(* Logix 5000 project; controller PLC_MCC1300_75F1 vendor 1 type 14 code 166 rev 32.11; software revision 32.04 *) (continued)
TYPE MAC_Conveyor_ALM :
STRUCT
   rgxStoppingFault : DINT[1];   // Generic stopping faults
   rgxFault : DINT[1];   // Generic faults
   rgxWarning : DINT[1];   // Generic warning
   rgxStoppingFault_M : DINT[2];   // Motor stopping faults
   rgxFault_M : DINT[2];   // Motor faults
   rgxWarning_M : DINT[2];   // Motor warning
   rgdFaultCode_M : DINT[2];   // Motor fault codes
END_STRUCT
END_TYPE

TYPE MAC_Conveyor_HMR :
STRUCT
   xSensorPresence1 : BOOL;   // Sensor presence 1 {x|x|x|x|O}
   xSensorPresence2 : BOOL;   // Sensor presence 2 {x|x|x|x|O}
   xSensorPresence3 : BOOL;   // Sensor presence 3 {x|x|x|x|O}
   xSensorPresence4 : BOOL;   // Sensor presence 4 {x|x|x|x|O}
   xSensorPresence5 : BOOL;   // Sensor presence 5 {x|x|x|x|O}
   xSensorPresence6 : BOOL;   // Sensor presence 6 {x|x|x|x|O}
   xHighPositionPopup1 : BOOL;   // High position popup {x|x|x|x|O}
   xLowPositionPopup1 : BOOL;   // Low position popup {x|x|x|x|O}
   xHighPositionPopup2 : BOOL;   // High position popup {x|x|x|x|O}
   xLowPositionPopup2 : BOOL;   // Low position popup {x|x|x|x|O}
   xHighPositionSquaring1 : BOOL;   // High position squaring {x|x|x|x|O}
   xLowPositionSquaring1 : BOOL;   // Low position squaring {x|x|x|x|O}
   xHighPositionSquaring2 : BOOL;   // High position squaring {x|x|x|x|O}
   xLowPositionSquaring2 : BOOL;   // Low position squaring {x|x|x|x|O}
   xCleaningEnabled : BOOL;   // Cleaning enabled {x|x|x|x|O}
   xWritingEnabled : BOOL;   // Writing enabled {x|x|x|x|O}
   xManualCommandEnabled : BOOL;   // Manual commands enabled {x|x|x|x|O}
   xVirtualDoorEnabled : BOOL;   // Virtual door enabled {x|x|x|x|O}
   xAuxFunctionEnabled : BOOL;   // Auxiliary function enabled {x|x|x|x|O}
   xIdPlatePresence : BOOL;   // Id plate presence {x|x|x|x|O}
   dState1 : DINT;   // State 1 (1=No anomaly, 3=Run, 7=Anomaly) {x|x|x|x|O}
   dState2 : DINT;   // State 2 (1=No anomaly, 3=Run, 7=Anomaly) {x|x|x|x|O}
   dState3 : DINT;   // State 3 (1=No anomaly, 3=Run, 7=Anomaly) {x|x|x|x|O}
   dState4 : DINT;   // State 4 (1=No anomaly, 3=Run, 7=Anomaly) {x|x|x|x|O}
   dStateSensor1 : DINT;   // State sensor 1 (1=No alarm, 7=Alarm) {x|x|x|x|O}
   dStateSensor2 : DINT;   // State sensor 2 (1=No alarm, 7=Alarm) {x|x|x|x|O}
   dStateSensor3 : DINT;   // State sensor 3(1=No alarm, 7=Alarm) {x|x|x|x|O}
   dStateSensor4 : DINT;   // State sensor 4(1=No alarm, 7=Alarm) {x|x|x|x|O}
   dStateSensor5 : DINT;   // State sensor 5(1=No alarm, 7=Alarm) {x|x|x|x|O}
   dStateSensor6 : DINT;   // State sensor 6(1=No alarm, 7=Alarm) {x|x|x|x|O}
   dErrorCode1 : DINT;   // Error code {x|x|x|x|O}
   dErrorCode2 : DINT;   // Error code {x|x|x|x|O}
   dErrorCode3 : DINT;   // Error code {x|x|x|x|O}
   dErrorCode4 : DINT;   // Error code {x|x|x|x|O}
   rgxMan : DINT;   // Manual commands {x|x|x|x|O}
END_STRUCT
END_TYPE

TYPE MAC_Conveyor_HMW :
STRUCT
   xLocalCleaningRequest : BOOL;   // Local cleaning request {x|x|x|x|O}
   xStopLocalCleaningRequest : BOOL;   // Stop local cleaning request {x|x|x|x|O}
   xEnableDisableManualCommand : BOOL;   // Enable/Disable manual commands {x|x|x|x|O}
   xSendDataToPLC : BOOL;   // Send plate data to PLC {x|x|x|x|O}
   xEnableDisableVirtualDoor : BOOL;   // Enable/Disable virtual door {x|x|x|x|O}
   xEnableDisableAuxFunction : BOOL;   // Enable/Disable auxiliary function {x|x|x|x|O}
   dParam_1_cmm : DINT;   // Auxiliary parameter 1 [mm/100] {mm/100|mm|x|x|O}
   dParam_2_cmm : DINT;   // Auxiliary parameter 2 [mm/100] {mm/100|mm|x|x|O}
   dParam_3_cmm : DINT;   // Auxiliary parameter 3 [mm/100] {mm/100|mm|x|x|O}
   dParam_4_cmm : DINT;   // Auxiliary parameter 4 [mm/100] {mm/100|mm|x|x|O}
   dParam_5_ms : DINT;   // Auxiliary parameter 5 [ms] {ms|ms|x|x|O}
   dParam_6_ms : DINT;   // Auxiliary parameter 6 [ms] {ms|ms|x|x|O}
   dParam_7_ms : DINT;   // Auxiliary parameter 7 [ms] {ms|ms|x|x|O}
   dParam_8_ms : DINT;   // Auxiliary parameter 8 [ms] {ms|ms|x|x|O}
   rgxMan : DINT;   // Manual commands {x|x|x|x|O}
END_STRUCT
END_TYPE

TYPE MAC_Conveyor_Single :
STRUCT
   ST_xInitialConditionOK : BOOL;   // Initial condition OK
   ST_xInitialConditionOK_BW : BOOL;   // Initial condition OK backward
   ST_xCleaningConditionOK : BOOL;   // Cleaning condition OK
   ST_xCleaningAccepted : BOOL;   // Cleaning accepted
   ST_xReqCleaning : BOOL;   // Request cleaning
   ST_xPlatePresence : BOOL;   // Plate presence memory
   ST_xPhasesInProgress : BOOL;   // Phases in progress
   ST_xCycleLoadUnload : BOOL;   // Cycle load/unload simultaneously
   ST_xStopMachineFault : BOOL;   // Stopped machine fault
   ST_xStopNextCycleFault : BOOL;   // Stop next cycle fault
   ST_xConditionOKStopCycle : BOOL;   // Condition OK for stop cycle
   ST_xOutputEnable : BOOL;   // Output enable
   ST_xMachineAlarm : BOOL;   // Machine alarm
   ST_xMachineWarning : BOOL;   // Machine warning
   ST_xIdPlatePresence : BOOL;   // Id plate presence
   ST_xFeedbackRotation : BOOL;   // Feedback rotation
   ST_xRampInProgress : BOOL;   // Ramp in progress
   ST_xAccInProgress : BOOL;   // Acceleration in progress
   ST_xDecInProgress : BOOL;   // Deceleration in progress
   ST_xWaitStopNextMachine : BOOL;   // Wait stop next machine
   ST_xWaitMachineStop : BOOL;   // Wait machine stop
   ST_xWaitReadyToMove : BOOL;   // Wait ready to move
   ST_xEnableControlError : BOOL;   // Enable control error
   ST_xManualMode : BOOL;   // Manual mode enabled
   ST_xPlateSynchronized : BOOL;   // Plate synchronized
   ST_xVirtualDoorEnabled : BOOL;   // Virtual door enabled
   ST_xDisableLoadUnloadOnStop : BOOL;   // Temporary disable of load/unload continuosly after a bit wait machine stop
   ST_xPlatePassageUpstream_FW : BOOL;   // Plate in passage upstream
   ST_xPlatePassageUpstream_BKW : BOOL;   // Plate in passage upstream
   ST_xPlatePassageDownstream_FW : BOOL;   // Plate in passage downstream
   ST_xPlatePassageDownstream_BKW : BOOL;   // Plate in passage downstream
   ST_xAxleReadyToMoveDelayed : BOOL;   // Axle ready to move delayed (NU)
   ST_xSafetyMovement : BOOL;   // Safety Mouvement
   ST_xReqDescent : BOOL;   // popup conveyor
   ST_xPhaseError : BOOL;   // Phase error, send lites to cullet
   ST_xAux1 : BOOL;   // ST Aux 1
   ST_xAux2 : BOOL;   // ST Aux 2
   ST_xAux3 : BOOL;   // ST Aux 3
   ST_xAux4 : BOOL;   // ST Aux 4
   OSR_xUnload : BOOL;   // OSR Unload
   OSR_xSynchroPhotocellHead : BOOL;   // OSR Synchronization photocell head
   OSR_xSynchroPhotocellTail : BOOL;   // OSR Synchronization photocell tail
   OSR_xPosReq : BOOL;   // OSR Positioning request
   OS_xLoad_FW : BOOL;   // OS Load forward
   OS_xUnload_FW : BOOL;   // OS Unload forward
   OS_xLoad_BW : BOOL;   // OS Load backward
   OS_xUnload_BW : BOOL;   // OS Unload backward
   OS_xUnpack : BOOL;   // OS Unpack convoy
   OS_xSynchroPhotocellHead : BOOL;   // OS Synchronization photocell head
   OS_xSynchroPhotocellTail : BOOL;   // OS Synchronization photocell tail
   OS_xChangeSpeed : BOOL;   // OS Dynamic change speed
   PH_x : DINT;   // Phases
   INPUT_xSyncroPhotocell_1 : BOOL;   // Sincro photocell / start count
   INPUT_xSyncroPhotocell_2 : BOOL;   // Sincro photocell / start count
   INPUT_xSquaringPhotocell_1 : BOOL;   // Squaring photocell #1
   INPUT_xSquaringPhotocell_2 : BOOL;   // Squaring photocell #2
   INPUT_xSquaringPhotocell_3 : BOOL;   // Squaring photocell #3
   INPUT_xSquaringPhotocell_4 : BOOL;   // Squaring photocell #4
   INPUT_xHighPositionSquaring_1 : BOOL;   // High position squaring #1
   INPUT_xLowPositionSquaring_1 : BOOL;   // Low position squaring #1
   INPUT_xHighPositionSquaring_2 : BOOL;   // High position squaring #2
   INPUT_xLowPositionSquaring_2 : BOOL;   // Low position squaring #2
   INPUT_xHighPositionPopup_1 : BOOL;   // High position pop-up
   INPUT_xLowPositionPopup_1 : BOOL;   // Low position pop-up
   INPUT_xHighPositionPopup_2 : BOOL;   // High position pop-up
   INPUT_xLowPositionPopup_2 : BOOL;   // Low position pop-up
   INPUT_xBrakingResistor_M1 : BOOL;   // Braking resistor
   INPUT_xDriveError_M1 : BOOL;   // Drive error
   INPUT_xDriveFeedback_M1 : BOOL;   // Drive feedback
   INPUT_xDriveInhibit_M1 : BOOL;
   INPUT_xDriveReady_M1 : BOOL;
   INPUT_xLocalSafetySwitch_M1 : BOOL;   // Local safety switch
   INPUT_xMotorThermalProbe_M1 : BOOL;   // Motor thermal probe
   INPUT_xProtectionMotor_M1 : BOOL;   // Protection motor
   INPUT_xBrakingResistor_M2 : BOOL;   // Braking resistor
   INPUT_xDriveError_M2 : BOOL;   // Drive error
   INPUT_xDriveFeedback_M2 : BOOL;   // Drive feedback
   INPUT_xDriveInhibit_M2 : BOOL;
   INPUT_xDriveReady_M2 : BOOL;
   INPUT_xLocalSafetySwitch_M2 : BOOL;   // Local safety switch
   INPUT_xMotorThermalProbe_M2 : BOOL;   // Motor thermal probe
   INPUT_xProtectionMotor_M2 : BOOL;   // Protection motor
   INPUT_xBrakingResistor_M3 : BOOL;   // Braking resistor
   INPUT_xDriveError_M3 : BOOL;   // Drive error
   INPUT_xDriveFeedback_M3 : BOOL;   // Drive feedback
   INPUT_xDriveInhibit_M3 : BOOL;
   INPUT_xDriveReady_M3 : BOOL;
   INPUT_xLocalSafetySwitch_M3 : BOOL;   // Local safety switch
   INPUT_xMotorThermalProbe_M3 : BOOL;   // Motor thermal probe
   INPUT_xProtectionMotor_M3 : BOOL;   // Protection motor
   INPUT_xBrakingResistor_M4 : BOOL;   // Braking resistor
   INPUT_xDriveError_M4 : BOOL;   // Drive error
   INPUT_xDriveFeedback_M4 : BOOL;   // Drive feedback
   INPUT_xDriveInhibit_M4 : BOOL;
   INPUT_xDriveReady_M4 : BOOL;
   INPUT_xLocalSafetySwitch_M4 : BOOL;   // Local safety switch
   INPUT_xMotorThermalProbe_M4 : BOOL;   // Motor thermal probe
   INPUT_xProtectionMotor_M4 : BOOL;   // Protection motor
   INPUT_xProtectionLiftingFrame_1 : BOOL;   // Protection lifting frame
   INPUT_xProtectionLiftingFrame_2 : BOOL;   // Protection lifting frame
   INPUT_xFeedBackLiftingFrame_1 : BOOL;   // Feedback lifting frame
   INPUT_xFeedBackLiftingFrame_2 : BOOL;   // Feedback lifting frame
   INPUT_xProtectionFun_1 : BOOL;   // Protection fun
   INPUT_xProtectionFun_2 : BOOL;   // Protection fun
   INPUT_xFeedbackVentilation_1 : BOOL;   // Feedback ventilation
   INPUT_xFeedbackVentilation_2 : BOOL;   // Feedback ventilation
   OUTPUT_xRisePopup_1 : BOOL;   // Rise popup
   OUTPUT_xDescentPopup_1 : BOOL;   // Descent popup
   OUTPUT_xRisePopup_2 : BOOL;   // Rise popup
   OUTPUT_xDescentPopup_2 : BOOL;   // Descent popup
   OUTPUT_xRiseSquaring_1 : BOOL;   // Rise squaring #1
   OUTPUT_xDescentSquaring_1 : BOOL;   // Descent squaring #1
   OUTPUT_xRiseSquaring_2 : BOOL;   // Rise squaring #2
   OUTPUT_xDescentSquaring_2 : BOOL;   // Descent squaring #2
   OUTPUT_xDriveEnable_M1 : BOOL;   // Drive enable
   OUTPUT_xPositioning_M1 : BOOL;   // Positiong
   OUTPUT_xReverse_M1 : BOOL;   // Reserve
   OUTPUT_xRun_M1 : BOOL;   // Run
   OUTPUT_xDriveEnable_M2 : BOOL;   // Drive enable
   OUTPUT_xPositioning_M2 : BOOL;   // Positiong
   OUTPUT_xReverse_M2 : BOOL;   // Reserve
   OUTPUT_xRun_M2 : BOOL;   // Run
   OUTPUT_xDriveEnable_M3 : BOOL;   // Drive enable
   OUTPUT_xPositioning_M3 : BOOL;   // Positiong
   OUTPUT_xReverse_M3 : BOOL;   // Reserve
   OUTPUT_xRun_M3 : BOOL;   // Run
   OUTPUT_xDriveEnable_M4 : BOOL;   // Drive enable
   OUTPUT_xPositioning_M4 : BOOL;   // Positiong
   OUTPUT_xReverse_M4 : BOOL;   // Reserve
   OUTPUT_xRun_M4 : BOOL;   // Run
   OUTPUT_xFunCommand_1 : BOOL;   // Fun command
   OUTPUT_xFunCommand_2 : BOOL;   // Fun command
   AUX_dPresetStopLoad_cmm : DINT;   // Preset Stop Load position [mm/100]
   AUX_dPresetStopUnload_cmm : DINT;   // Preset Stop Unload position [mm/100]
   AUX_dAccSpace_cmm : DINT;   // Acceleration Space [mm/100]
   AUX_dDecSpace_cmm : DINT;   // Acceleration Space [mm/100]
   AUX_dReqSpeed_mm_min : DINT;   // Conveyor requested speed [mm/min]
   AUX_dAbsPosTarget_M1_cmm : DINT;   // Absolute positioning target [mm/100]
   AUX_dAbsPosTarget_M2_cmm : DINT;   // Absolute positioning target [mm/100]
   AUX_dAbsPosTarget_M3_cmm : DINT;   // Absolute positioning target [mm/100]
   AUX_dAbsPosTarget_M4_cmm : DINT;   // Absolute positioning target [mm/100]
   AUX_dPhPosTarget_cmm : DINT;   // Photocell positioning target [mm/100]
   AUX_dQtaLites : DINT;   // Qta lites on conveyor
   TmON_AxleReadyToMoveDelayed : TIMER;   // Axle ready to move delayed (NU)
   tmON_FeedbackTimeOut_M1 : TIMER;   // Feedback time out
   tmOF_DriveEnable_M1 : TIMER;   // Drive enable timer
   tmOF_PowerSaving_M1 : TIMER;   // Power saving timer
   tmON_FeedbackTimeOut_M2 : TIMER;   // Feedback time out
   tmOF_DriveEnable_M2 : TIMER;   // Drive enable timer
   tmOF_PowerSaving_M2 : TIMER;   // Power saving timer
   tmON_FeedbackTimeOut_M3 : TIMER;   // Feedback time out
   tmOF_DriveEnable_M3 : TIMER;   // Drive enable timer
   tmOF_PowerSaving_M3 : TIMER;   // Power saving timer
   tmON_FeedbackTimeOut_M4 : TIMER;   // Feedback time out
   tmOF_DriveEnable_M4 : TIMER;   // Drive enable timer
   tmOF_PowerSaving_M4 : TIMER;   // Power saving timer
   tmON_PosTimeOut_1 : TIMER;   // Positioning timeout 1
   tmON_PosTimeOut_2 : TIMER;   // Positioning timeout 2
   tmON_PosTimeOut_3 : TIMER;   // Positioning timeout 3
   tmON_Wait : TIMER;   // Wait for glass process
   tmON_AuxFunction1 : TIMER;   // Timer auxiliary function 1
   tmON_AuxFunction2 : TIMER;   // Timer auxiliary function 2
   tmON_AuxFunction3 : TIMER;   // Timer auxiliary function 3
   tmON_AuxFunction4 : TIMER;   // Timer auxiliary function 4
   tmON_AuxFunction5 : TIMER;   // Timer auxiliary function 5
   tmON_AuxFunction6 : TIMER;   // Timer auxiliary function 6
   tmON_AuxFunction7 : TIMER;   // Timer auxiliary function 7
   tmON_AuxFunction8 : TIMER;   // Timer auxiliary function 8
   tmON_AuxFunction9 : TIMER;   // Timer auxiliary function 9
   TmON : TIMER[16];
   tmOF_MCD_M1 : TIMER;
   tmOF_MCD_M2 : TIMER;
   tmOF_MCD_M3 : TIMER;
   tmOF_MCD_M4 : TIMER;
END_STRUCT
END_TYPE

TYPE MAC_Conveyor_ZC :
STRUCT
   CONST_dMachineNumb : DINT;   // Machine number [Mxxx = xxx*10]
   CONST_dMachineZoneNumb : DINT;   // Machine zones number [0 = No zones; 2 = 2 Zones; etc...]
   CONST_dMotorNumber : DINT;   // Number of motor [0 = Single motor; 2 = 2 motors; etc...]
   CONST_dOriginSetpoint_cmm : DINT;   // Distance from the beggining (From origin to split line) [mm/100]
   CONST_dPresetFeedbackTime_ms : DINT;   // Preset feedback time [ms]
   CONST_dPresetStopLoad_cmm : DINT;   // Preset stop load [mm/100]
   CONST_dConveyorLength_cmm : DINT;   // Conveyor length [mm/100]
   CONST_dConveyorWidth_cmm : DINT;   // Conveyor width [mm/100]
   CONST_dConveyorZones_cmm : DINT[6];   // [0]Zone1 [mm/100]; [1]Zone2 [mm/100]; etc...
   CONST_dSyncroPhPosition_cmm : DINT;   // Synchronization photocell position [mm/100]
   CONST_dSyncroPhWindow_cmm : DINT;   // Synchronization photocell window [mm/100]
   CONST_dMainRefSpeedIndx : DINT;   // Main reference speed [Index "RefSpeed"]
   CONST_xEnableSyncHead : BOOL;   // Enable synchronization on head
   CONST_xEnableSyncTail : BOOL;   // Enable synchronization on tail
   ST_xCleaningConditionOK : BOOL;   // Cleaning condition OK
   ST_xStopMachineFault : BOOL;   // Stopped machine faults
   ST_xStopNextCycleFault : BOOL;   // Stopped next cycle faults
   ST_xConditionOKStopCycle : BOOL;   // Condition OK for stop cycle
   ST_xManualMode : BOOL;   // Manual mode enabled
   ST_xOutputEnable : BOOL;   // Output enable
   ST_xMachineFault : BOOL;   // Machine with faults
   ST_xFeedbackRotation : BOOL;   // Feedback rotation
   ST_BrakeRelease : BOOL;   // Brake release
   ST_xRampInProgress : BOOL;   // Ramp in progress
   ST_xAccInProgress : BOOL;   // Acceleration in progress
   ST_xDecInProgress : BOOL;   // Deceleration in progress
   ST_xConveyorInRun : BOOL;   // Conveyor in run
   ST_ConveyorRunning : BOOL;   // Conveyor running
   ST_ConvoyInProgress : BOOL;   // Convoy transiting on conveyor
   ST_xStopConveyor : BOOL;   // Stop conveyor
   ST_xPlateInStopPos : BOOL;   // Plate in stop position
   ST_xPlateOnSplitLine : BOOL;   // Plate on split line downstream
   ST_xHeadPresence : BOOL;   // Head presence on conveyor
   ST_xTailPresence : BOOL;   // Tail presence on conveyor
   ST_xEnableControlError : BOOL;   // Enable control error
   ST_xPlateSynchronized : BOOL;   // Plate synchronized
   ST_xSinchroPhError : BOOL;   // Sinchronization error
   ST_xBypassSynchroAnomaly : BOOL;   // Bypass synchronization error
   OSR_xSynchroPhotocellHead : BOOL;   // OSR Synchronization photocell head
   OSR_xSynchroPhotocellTail : BOOL;   // OSR Synchronization photocell tail
   OSR_xStartCount : BOOL;   // OSR Start count positionig
   OSR_xEndSync : BOOL;   // OSR End synchronization
   OS_xSynchroPhotocellHead : BOOL;   // OS Synchronization photocell head
   OS_xSynchroPhotocellTail : BOOL;   // OS Synchronization photocell tail
   OS_xStartCount : BOOL;   // OS Start count positionig
   OS_xEndSync : BOOL;   // OS End synchronization
   PH : MAC_Conveyor_ZC_PH;   // Phases
   INPUT_xSyncroPhotocell : BOOL;   // Syncronization Photocell
   INPUT_xNextConveyorInRun : BOOL;   // Next conveyor in run
   INPUT_xBrakingResistor : DINT;   // Braking Resistor
   INPUT_xDriveInhibit : DINT;   // Drive inhibit
   INPUT_xDriveReady : DINT;   // Drive ready
   INPUT_xDriveError : DINT;   // Drive Error
   INPUT_xDriveFeedback : DINT;   // Drive Feedback
   INPUT_xDriveDeceleration : DINT;   // Drive deceleration
   INPUT_xLocalSafetySwitch : DINT;   // Local Safety Switch
   INPUT_xMotorThermalProbe : DINT;   // Motor Thermal Probe
   INPUT_xProtectionMotor : DINT;   // Protection Motor
   INPUT_xProtectionCoolingFan : DINT;   // Protection cooling fan
   INPUT_xFeedbackCoolingFan : DINT;   // Feedback cooling fan
   INPUT_xDrivePositionReached : DINT;   // Drive position reached
   INPUT_dRefSpeed_mm_min : DINT[3];   // Reference speed [0]Cleaning speed [mm/min]; [1] Lehr speed [mm/min]; [2] Automatic speed; etc...
   OUTPUT_xDriveReset : DINT;   // Drive reset faults
   OUTPUT_xDriveEnable : DINT;   // Output
   OUTPUT_xRun : DINT;   // Run
   OUTPUT_xReverse : DINT;   // Reverse
   OUTPUT_xPositioning : DINT;   // Positioning
   OUTPUT_xChangeSpeed : DINT;   // Change speed
   AUX_dCountFeedbackTime_ms : DINT;   // Counter feedback time [ms]
   AUX_dReqTarget_cmm : DINT;   // Request target for positioning [mm/100]
   AUX_dReqSpeed_mm_min : DINT[2];   // Conveyor requested speed [mm/min]
   AUX_dRealSpeed_mm_min : DINT[2];   // Conveyor real speed [mm/min]
   AUX_dHeadPosition_cmm : DINT;   // Plate head position [mm/100]
   AUX_dTailPosition_cmm : DINT;   // Plate tail position [mm/100]
   AUX_dAccSpace_cmm : DINT;   // Acceleration space [mm/100]
   AUX_dDecSpace_cmm : DINT;   // Deceleration space [mm/100]
   AUX_dLastIDPlateLoaded : DINT;   // Last ID plate loaded
   AUX_rAcceleration_m_s2 : REAL;   // Acceleration ramp [m/s2]
   AUX_rDeceleration_m_s2 : REAL;   // Deceleration ramp [m/s2]
   AUX_rSpeedIncrement_mm_min : REAL[2];   // Speed increment [mm/min]
   AUX_rStepAdvancement : REAL[2];   // Step advancement [mm/10 per Scan]
   AUX_rHeadPosition_cmm : REAL;   // Head position [mm/100]
   AUX_rTailPosition_cmm : REAL;   // Tail position [mm/100]
   tmON_FeedbackTimeOut : TIMER[2];   // Feedback time out
   tmOF_DriveEnable : TIMER[2];   // Drive enable timer
   tmON_Wait : TIMER;   // Wait for glass process
   tmON_SyncTimeout : TIMER;   // Time out synchronization photocell
   tmOF_SyncTimeout : TIMER;   // Time out synchronization photocell
   tmON_PhFilter : TIMER;   // Start count photocell filter
END_STRUCT
END_TYPE

TYPE MAC_Conveyor_ZC_ALM :
STRUCT
   rgxStoppingFault : MAC_Conveyor_ZC_ALM_SF[1];   // Generic stopping faults
   rgxFault : MAC_Conveyor_ZC_ALM_F[1];   // Generic faults
   rgxWarning : MAC_Conveyor_ZC_ALM_W[1];   // Generic warning
   rgxStoppingFault_M : MAC_Conveyor_ZC_ALM_SFM[2];   // Motor stopping faults
   rgxFault_M : MAC_Conveyor_ZC_ALM_FM[2];   // Motor faults
   rgxWarning_M : MAC_Conveyor_ZC_ALM_WM[2];   // Motor warning
   rgdFaultCode_M : DINT[2];   // Motor fault codes
END_STRUCT
END_TYPE

TYPE MAC_Conveyor_ZC_ALM_F :
STRUCT
   x0 : BOOL;
   x1 : BOOL;
   x2 : BOOL;
   x3 : BOOL;
   x4 : BOOL;
   x5 : BOOL;
   x6 : BOOL;
   x7 : BOOL;
   x8 : BOOL;
   x9 : BOOL;
   x10 : BOOL;
   x11 : BOOL;
   x12 : BOOL;
   x13 : BOOL;
   x14 : BOOL;
   x15 : BOOL;
   x16 : BOOL;
   x17 : BOOL;
   x18 : BOOL;
   x19 : BOOL;
   x20 : BOOL;
   x21 : BOOL;
   x22 : BOOL;
   x23 : BOOL;
   x24 : BOOL;
   x25 : BOOL;
   x26 : BOOL;
   x27 : BOOL;
   x28 : BOOL;
   x29 : BOOL;
   x30 : BOOL;
   x31 : BOOL;
END_STRUCT
END_TYPE

TYPE MAC_Conveyor_ZC_ALM_FM :
STRUCT
   x0 : BOOL;   // Protection cooling fan
   x1 : BOOL;
   x2 : BOOL;
   x3 : BOOL;
   x4 : BOOL;
   x5 : BOOL;
   x6 : BOOL;
   x7 : BOOL;
   x8 : BOOL;
   x9 : BOOL;
   x10 : BOOL;
   x11 : BOOL;
   x12 : BOOL;
   x13 : BOOL;
   x14 : BOOL;
   x15 : BOOL;
   x16 : BOOL;
   x17 : BOOL;
   x18 : BOOL;
   x19 : BOOL;
   x20 : BOOL;
   x21 : BOOL;
   x22 : BOOL;
   x23 : BOOL;
   x24 : BOOL;
   x25 : BOOL;
   x26 : BOOL;
   x27 : BOOL;
   x28 : BOOL;
   x29 : BOOL;
   x30 : BOOL;
   x31 : BOOL;
END_STRUCT
END_TYPE

TYPE MAC_Conveyor_ZC_ALM_SF :
STRUCT
   x0 : BOOL;
   x1 : BOOL;
   x2 : BOOL;
   x3 : BOOL;
   x4 : BOOL;
   x5 : BOOL;
   x6 : BOOL;
   x7 : BOOL;
   x8 : BOOL;
   x9 : BOOL;
   x10 : BOOL;
   x11 : BOOL;
   x12 : BOOL;
   x13 : BOOL;
   x14 : BOOL;
   x15 : BOOL;
   x16 : BOOL;
   x17 : BOOL;
   x18 : BOOL;
   x19 : BOOL;
   x20 : BOOL;
   x21 : BOOL;
   x22 : BOOL;
   x23 : BOOL;
   x24 : BOOL;
   x25 : BOOL;
   x26 : BOOL;
   x27 : BOOL;
   x28 : BOOL;
   x29 : BOOL;
   x30 : BOOL;
   x31 : BOOL;
END_STRUCT
END_TYPE

TYPE MAC_Conveyor_ZC_ALM_SFM :
STRUCT
   x0 : BOOL;   // Protection motor
   x1 : BOOL;   // Drive error
   x2 : BOOL;   // Drive feedback error
   x3 : BOOL;   // Local safety switch
   x4 : BOOL;   // Motor thermal probe
   x5 : BOOL;   // Braking resistor fault
   x6 : BOOL;
   x7 : BOOL;
   x8 : BOOL;
   x9 : BOOL;
   x10 : BOOL;
   x11 : BOOL;
   x12 : BOOL;
   x13 : BOOL;
   x14 : BOOL;
   x15 : BOOL;
   x16 : BOOL;
   x17 : BOOL;
   x18 : BOOL;
   x19 : BOOL;
   x20 : BOOL;
   x21 : BOOL;
   x22 : BOOL;
   x23 : BOOL;
   x24 : BOOL;
   x25 : BOOL;
   x26 : BOOL;
   x27 : BOOL;
   x28 : BOOL;
   x29 : BOOL;
   x30 : BOOL;
   x31 : BOOL;
END_STRUCT
END_TYPE

TYPE MAC_Conveyor_ZC_ALM_W :
STRUCT
   x0 : BOOL;   // Plate not synchronized
   x1 : BOOL;
   x2 : BOOL;
   x3 : BOOL;
   x4 : BOOL;
   x5 : BOOL;
   x6 : BOOL;
   x7 : BOOL;
   x8 : BOOL;
   x9 : BOOL;
   x10 : BOOL;
   x11 : BOOL;
   x12 : BOOL;
   x13 : BOOL;
   x14 : BOOL;
   x15 : BOOL;
   x16 : BOOL;
   x17 : BOOL;
   x18 : BOOL;
   x19 : BOOL;
   x20 : BOOL;
   x21 : BOOL;
   x22 : BOOL;
   x23 : BOOL;
   x24 : BOOL;
   x25 : BOOL;
   x26 : BOOL;
   x27 : BOOL;
   x28 : BOOL;
   x29 : BOOL;
   x30 : BOOL;
   x31 : BOOL;
END_STRUCT
END_TYPE

TYPE MAC_Conveyor_ZC_ALM_WM :
STRUCT
   x0 : BOOL;
   x1 : BOOL;
   x2 : BOOL;
   x3 : BOOL;
   x4 : BOOL;
   x5 : BOOL;
   x6 : BOOL;
   x7 : BOOL;
   x8 : BOOL;
   x9 : BOOL;
   x10 : BOOL;
   x11 : BOOL;
   x12 : BOOL;
   x13 : BOOL;
   x14 : BOOL;
   x15 : BOOL;
   x16 : BOOL;
   x17 : BOOL;
   x18 : BOOL;
   x19 : BOOL;
   x20 : BOOL;
   x21 : BOOL;
   x22 : BOOL;
   x23 : BOOL;
   x24 : BOOL;
   x25 : BOOL;
   x26 : BOOL;
   x27 : BOOL;
   x28 : BOOL;
   x29 : BOOL;
   x30 : BOOL;
   x31 : BOOL;
END_STRUCT
END_TYPE

TYPE MAC_Conveyor_ZC_HMR :
STRUCT
   xManualCommandEnabled : BOOL;   // Manual commands enabled {x|x|x|x|O}
   xCleaningEnabled : BOOL;   // Cleaning enabled {x|x|x|x|O}
   xPlatePresence : BOOL;   // Plate present {x|x|x|x|O}
   rgdState : DINT[2];   // State (1=No anomaly, 3=Run, 7=Anomaly) {x|x|x|x|O}
   rgxMan : MAC_Conveyor_ZC_HMWR_Man;   // Manual commands {x|x|x|x|O}
END_STRUCT
END_TYPE

TYPE MAC_Conveyor_ZC_HMW :
STRUCT
   xLocalCleaningRequest : BOOL;   // Local cleaning request {x|x|x|x|O}
   xEnableDisableManualCommand : BOOL;   // Enable / Disable manual commands {x|x|x|x|O}
   rgxMan : MAC_Conveyor_ZC_HMWR_Man;   // Manual commands {x|x|x|x|O}
END_STRUCT
END_TYPE

TYPE MAC_Conveyor_ZC_HMWR_Man :
STRUCT
   xCmdFwd : INT;   // Run forward
   xCmdBwd : INT;   // Run backward
   xAllFwd : BOOL;   // Run all forward
   xAllBwd : BOOL;   // Run all backward
END_STRUCT
END_TYPE

TYPE MAC_Conveyor_ZC_IN_MOTION :
STRUCT
   DR_MAJ_M : MOTION_INSTRUCTION[2];   // Drive jog
   DR_MAM_M : MOTION_INSTRUCTION[2];   // Drive positioning
   DR_MRP_M : MOTION_INSTRUCTION[2];   // Drive reset count
   DR_MAR_M : MOTION_INSTRUCTION[2];   // Drive registration
   DR_MASall_M : MOTION_INSTRUCTION[2];   // Drive stop
   DR_MASjog_M : MOTION_INSTRUCTION[2];   // Drive stop
   DR_MASpos_M : MOTION_INSTRUCTION[2];   // Drive stop
END_STRUCT
END_TYPE

TYPE MAC_Conveyor_ZC_OUT_MOTION :
STRUCT
   DR_MSO_M : MOTION_INSTRUCTION[2];   // Drive ON
   DR_MSF_M : MOTION_INSTRUCTION[2];   // Drive OFF
   DR_MASR_M : MOTION_INSTRUCTION[2];   // Drive reset faults
   DR_MAJ_M : MOTION_INSTRUCTION[2];   // Drive jog
   DR_MAM_M : MOTION_INSTRUCTION[2];   // Drive positioning
   DR_MAG_M : MOTION_INSTRUCTION[2];   // Drive gearing
   DR_MRP_M : MOTION_INSTRUCTION[2];   // Drive reset count
   DR_MAR_M : MOTION_INSTRUCTION[2];   // Drive enable registration
   DR_MDR_M : MOTION_INSTRUCTION[2];   // Drive disable registration
   DR_MCD_M : MOTION_INSTRUCTION[2];   // Drive change speed
   DR_MASall_M : MOTION_INSTRUCTION[2];   // Drive stop
   DR_MASjog_M : MOTION_INSTRUCTION[2];   // Drive stop
   DR_MASpos_M : MOTION_INSTRUCTION[2];   // Drive stop
END_STRUCT
END_TYPE

TYPE MAC_Conveyor_ZC_PH :
STRUCT
   x : SINT;   // Acceleration
   x8 : BOOL;   // Acceleration all
   x9 : BOOL;
   x10 : BOOL;
   x11 : BOOL;   // Stop conveyor forseen from external management
   x12 : BOOL;   // Bypass stop conveyor
   x13 : BOOL;   // Stop forseen for Pick-up
   x14 : BOOL;   // Positioning request
   x15 : BOOL;   // Stop conveyor request
   x16 : BOOL;   // Synchronization in progress
   x17 : BOOL;   // Synchronization error
   x18 : BOOL;
   x19 : BOOL;
   x20 : BOOL;
   x21 : BOOL;   // End stop/position request
   x22 : BOOL;
   x23 : BOOL;
   x24 : BOOL;   // Pick-up plate from conveyor in progress
   x25 : BOOL;
   x26 : BOOL;
   x27 : BOOL;
   x28 : BOOL;
   x29 : BOOL;
   x30 : BOOL;
   x31 : BOOL;
END_STRUCT
END_TYPE

TYPE MAC_Popup_ZC :
STRUCT
   ST_xTunnelType : BOOL;   // Tunnel type popup
   ST_xConditionToUnload : BOOL;   // Condition OK for unload
   ST_xCleaningConditionOK : BOOL;   // Cleaning condition OK
   ST_xCleaningAccepted : BOOL;   // Cleaning accepted
   ST_xReqCleaning : BOOL;   // Cleaning request
   ST_xStopMachineFault : BOOL;   // Stopped machine faults
   ST_xStopNextCycleFault : BOOL;   // Stopped next cycle faults
   ST_xConditionOKForStopCycle : BOOL;   // Condition OK for stop cycle
   ST_xManualMode : BOOL;   // Manual mode enabled
   ST_xOutputEnable : BOOL;   // Output enable
   ST_xMachineEmergencyAlarm : BOOL;   // Machine with emergency alarm
   ST_xMachineAlarm : BOOL;   // Machine with faults
   ST_xMachineWarning : BOOL;   // Machine with warning
   ST_xInitialConditionForRise : BOOL;   // Initial condition for rise popup
   ST_xInitialConditionForDescend : BOOL;   // Initial condition for descend popup
   ST_xRequestRise : BOOL;   // Request rise popup
   ST_xRequestDescend : BOOL;   // Request descend popup
   ST_xExternalConditionToRise : BOOL;   // External condition to rise popup
   ST_xExternalConditionToDescend : BOOL;   // External condition to descend popup
   ST_xOutOfEncumbrance : BOOL;   // Popup out of encumbrance
   ST_xPlatePresence : BOOL;   // Popup plate presence (Plate Data on Belts (side leg))
   ST_xConditionToReceiveGlass : BOOL;   // Popup condition to receive glass
   ST_xConditionForUpperConveyor : BOOL;   // Popup condition for upper conveyor
   ST_xFeedbackRotation : BOOL;   // Feedback rotation
   ST_xRampInProgress : BOOL;   // Ramp in progress
   ST_xAccInProgress : BOOL;   // Acceleration in progress
   ST_xDecInProgress : BOOL;   // Deceleration in progress
   ST_xPlateInStopPos : BOOL;   // Plate in stop position on conveyor
   ST_xHeadPresence : BOOL;   // Head presence on conveyor
   ST_xTailPresence : BOOL;   // Tail presence on conveyor
   ST_xEnableControlError : BOOL;   // Enable control error
   ST_xPlatePresentOnPopup : BOOL;   // Plate present on popup (Plate Data on Main Line)
   ST_xPlateToBeUnload : BOOL;   // Plate to be unload
   ST_xPlateToBeUnloadOpSide : BOOL;   // Plate to be unload to operator side
   ST_xPlateToBeUnloadOppOpSide : BOOL;   // Plate to be unload to opposite operator side
   ST_xPlateUnderPopup : BOOL;   // Plate under popup
   ST_xPlateToStopAfterPos : BOOL;   // Plate presence to stop after positioning
   ST_xPopupChangeDest : BOOL;   // Popup change destination
   ST_xPhasesInProgress : BOOL;   // Phases in progress
   ST_xPlateDataReadyToSend : BOOL;   // Plate data ready to send
   ST_xPlateDataSentToSideLeg : BOOL;   // Plate data sent to side leg
   ST_xPlateRemovedBySideLeg : BOOL;   // Plate removed by side leg
   ST_xPlateLoadedBySideLeg : BOOL;   // Plate loaded by side leg
   ST_xIndexConsPositioning : BOOL;   // Index consistance positioning
   ST_xPlateComingToPopup : BOOL;   // Plate coming is destinated to popup
   ST_xPlateStopToPopup : BOOL;   // Plate stop is destinated to popup
   ST_xPlateToBothComing : BOOL;   // Plate coming is destinated to both sides popup
   ST_xPlateToSingleComing : BOOL;   // Plate coming is destinated only to this section of pupup
   ST_xConvoyComing : BOOL;   // Plate coming is a convoy (to both sides of popup)
   ST_xPlateToBothPositioning : BOOL;   // Plate positioning is destinated to both sides popup
   ST_xPlateToSinglePositioning : BOOL;   // Plate positioning is destinated only to this section of pupup
   ST_xConvoyPositioning : BOOL;   // Plate positioning is a convoy (to both sides of popup)
   ST_xStopPreviousConveyor : BOOL;   // Stop previous conveyor
   ST_xConditionToStopPrevious : BOOL;   // Condition to stop previous conveyor
   ST_xSaturationConditionPopup : BOOL;   // Saturation condition on popup
   ST_xSaturationConditionPrevious : BOOL;   // Saturation condition on previous conveyor
   ST_xSaturationConditionThis : BOOL;   // Saturation condition on this conveyor
   ST_xPrevConvFreeAfterPos : BOOL;   // Previous conveyor free after positioning plate
   ST_xConvFreeForPos : BOOL;   // Conveyor free for positioning
   ST_xPlateInPositionToRise : BOOL;   // Plate in position to rise
   PH_xRise : BOOL;   // Rise phase
   PH_xEndRise : BOOL;   // End rise phase
   PH_xDescend : BOOL;   // Descend phase
   PH_xEndDescend : BOOL;   // End descend phase
   OS_xStartPositioning : BOOL;   // OS Start positioning
   OS_xTimeoutPositioning : BOOL;   // OS Timeout positioning
   OS_xPlateDataSentToSideLeg : BOOL;   // OS Plate data sent to side leg
   OS_xPlateRemovedBySideLeg : BOOL;   // OS Plate removed by side leg
   OS_xPlateLoadedBySideLeg : BOOL;   // OS Plate loaded by side leg
   OS_xSaturationOnPopup : BOOL;   // OS Saturation on popup
   OS_xSaturationOnPrevious : BOOL;   // OS Saturation on previous conveyor
   OS_xSaturationOnThis : BOOL;   // OS Saturation on this conveyor
   OS_xLastFreeForPos : BOOL;   // OS Last conveyor free for positioning
   OS_xChangeDestAfterRestart : BOOL;   // OS Change dest after restart because positioning impossible
   OS_xChangeDestAfterPopup : BOOL;   // OS Change dest after popup (undertaker function)
   OSR_xChangeDestAfterPopup : BOOL;   // OSR Change dest after popup (undertaker function)
   OS : DINT;   // OS (spare)
   PH_x : DINT;   // Phases (spare)
   INPUT_xLiftingProtectionMotor : BOOL;   // Lifting protection motor
   INPUT_xLiftingFeedbackMotor : BOOL;   // Lifting feedback motor
   INPUT_xLiftingSafetySwitch : BOOL;   // Lifting Local Safety Switch
   INPUT_xProtectionCoolingFan : BOOL;   // Cooling fan protection
   INPUT_xFeedbackCoolingFan : BOOL;   // Cooling fan protection
   INPUT_xPopupHigh : BOOL;   // Popup in high feedback
   INPUT_xPopupLow : BOOL;   // Popup in low position
   INPUT_xBrakingResistor : BOOL;   // Braking Resistor
   INPUT_xDriveInhibit : BOOL;   // Drive inhibit
   INPUT_xDriveReady : BOOL;   // Drive ready
   INPUT_xDriveError : BOOL;   // Drive Error
   INPUT_xDriveFeedback : BOOL;   // Drive Feedback
   INPUT_xBeltsSafetySwitch : BOOL;   // Belts Local Safety Switch
   INPUT_xBeltsMotorThermalProbe : BOOL;   // Belts Motor Thermal Probe
   INPUT_xBeltsProtectionMotor : BOOL;   // Belts Protection Motor
   INPUT_xConveyorOpSideInRun : BOOL;   // Conveyor in run operator side
   INPUT_xConveyorOppOpSideInRun : BOOL;   // Conveyor in run opposite operator side
   INPUT_dRefSpeed_mm_min : DINT;   // Reference speed [mm/min]
   OUTPUT_xPopupLifting : BOOL;   // Popup lifting
   OUTPUT_xPopupDescent : BOOL;   // Popup descent
   OUTPUT_xPopupVentilation : BOOL;   // Popup ventilation
   OUTPUT_xDriveReset : BOOL;   // Drive reset faults
   OUTPUT_xDriveEnable : BOOL;   // Output
   OUTPUT_xRun : BOOL;   // Run
   OUTPUT_xReverse : BOOL;   // Reverse
   OUTPUT_xPositioning : BOOL;   // Positioning
   OUTPUT_xChangeSpeed : BOOL;   // Change speed
   AUX_dStartPosition_cmm : DINT;   // Distance from the beggining (From origin to split line) [mm/100]
   AUX_dEndPosition_cmm : DINT;   // Distance from the end (From origin to split line) [mm/100]
   AUX_dPresetFeedbackTime_ms : DINT;   // Preset feedback time [ms]
   AUX_dPresetStopLoad_cmm : DINT;   // Preset stop load [mm/100]
   AUX_dSpeedConveyor_mm_min : DINT;   // Conveyor speed [mm/min]
   AUX_dPopupLength_cmm : DINT;   // Popup length [mm/100]
   AUX_dReactionTime_ms : DINT;   // Reaction time [ms]
   AUX_dWindowSearch_cmm : DINT;   // Window search length [mm/100]
   AUX_dChangeCulletReasonIndex : DINT;   // Change destination to cullet reason index [Num]
   AUX_dDestMaskOpSide : DINT;   // Destination available on sideleg to operator side (If 0 = no destinations) [Num]
   AUX_dDestMaskOppOpSide : DINT;   // Destination available on sideleg to opposite operator side (If 0 = no destinations) [Num]
   AUX_dCountFeedbackTime_ms : DINT;   // Counter feedback time [ms]
   AUX_dReqTarget_cmm : DINT;   // Request target for positioning [mm/100]
   AUX_dPosition_cmm : DINT;   // Plate position [mm/100]
   AUX_dStartPosWithReaction_cmm : DINT;   // Plate position start search [mm/100]
   AUX_dPosPhotocell_cmm : DINT;   // Positioning photocell position [mm/100]
   AUX_dIndexHead : DINT;   // Index head for positioning
   AUX_dIndexTail : DINT;   // Index tail for positioning
   AUX_dPosTimeout : DINT;   // Positioning timeout space
   AUX_dIndexPlateStop : DINT;   // Index of plate to stop on popup
   AUX_dIndexPositioning : DINT;   // Index of plate to position
   AUX_dMemoryPositioning : DINT;   // Index memory of plate to position
   AUX_dIndexPlatePositioned : DINT;   // Index of plate positioned
   AUX_dIndexPlateFree : DINT;   // Index of plate to position
   AUX_dLastIndexFreeForPos : DINT;   // Index of last plate free for positioning
   AUX_dIndexPlateToChangeDestAfterPopup : DINT;   // Index of plate to change destination after popup (undertaker function)
   AUX_tSearchPlateData : UDT_SearchPlateAuxData;   // Auxiliary data for searching plate
   tSearchPlateFree : GP_TrackingSearchPlate_STC;   // Data for search plate under popup
   tSearchPlateStop : GP_TrackingSearchPlate_STC;   // Data for search plate stop on popup
   tSearchPlateChangeDestAfterPopup : GP_TrackingSearchPlate_STC;   // Data for search plate to change destination after popup
   tmON_LiftingTimeOut : TIMER;   // Lifting time out
   tmON_LiftingFeedbackTimeOut : TIMER;   // Lifting Feedback time out
   tmOF_DriveEnable : TIMER;   // Drive enable timer
   tmOF_WaitBothEndLift : TIMER;   // Wait end lift of both popup
   tmOF_Wait : TIMER;   // Wait end phases of popup
   tmON_Saturation : TIMER;   // Saturation timer
   tmON_ReentryPlate : TIMER;   // Reentry plate timer
   tmON_Positioning : TIMER;   // Positioning timer
END_STRUCT
END_TYPE
